   // hmiStns[1].wip[18].pnCode[6] := 1000;
   // hmiStns[1].wip[18].pnCode[7] := 1000;
   // hmiStns[1].wip[19].pnCode[0] := 1000;
   // hmiStns[1].wip[19].pnCode[1] := 1000;
   // hmiStns[1].wip[19].pnCode[2] := 1000;
   // hmiStns[1].wip[19].pnCode[3] := 1000;
   // hmiStns[1].wip[19].pnCode[4] := 1000;
   // hmiStns[1].wip[19].pnCode[5] := 1000;
   // hmiStns[1].wip[19].pnCode[6] := 1000;
   // hmiStns[1].wip[19].pnCode[7] := 1000;
   // hmiStns[1].wip[20].pnCode[0] := 1000;
   // hmiStns[1].wip[20].pnCode[1] := 1000;
   // hmiStns[1].wip[20].pnCode[2] := 1000;
   // hmiStns[1].wip[20].pnCode[3] := 1000;
   // hmiStns[1].wip[20].pnCode[4] := 1000;
   // hmiStns[1].wip[20].pnCode[5] := 1000;
   // hmiStns[1].wip[20].pnCode[6] := 1000;
   // hmiStns[1].wip[20].pnCode[7] := 1000;
   // hmiStns[1].wip[21].pnCode[0] := 1000;
   // hmiStns[1].wip[21].pnCode[1] := 1000;
   // hmiStns[1].wip[21].pnCode[2] := 1000;
   // hmiStns[1].wip[21].pnCode[3] := 1000;
   // hmiStns[1].wip[21].pnCode[4] := 1000;
   // hmiStns[1].wip[21].pnCode[5] := 1000;
   // hmiStns[1].wip[21].pnCode[6] := 1000;
   // hmiStns[1].wip[21].pnCode[7] := 1000;
   // hmiStns[1].wip[22].pnCode[0] := 1000;
   // hmiStns[1].wip[22].pnCode[1] := 1000;
   // hmiStns[1].wip[22].pnCode[2] := 1000;
   // hmiStns[1].wip[22].pnCode[3] := 1000;
   // hmiStns[1].wip[22].pnCode[4] := 1000;
   // hmiStns[1].wip[22].pnCode[5] := 1000;
   // hmiStns[1].wip[22].pnCode[6] := 1000;
   // hmiStns[1].wip[22].pnCode[7] := 1000;
   // hmiStns[1].wip[23].pnCode[0] := 1000;
   // hmiStns[1].wip[23].pnCode[1] := 1000;
   // hmiStns[1].wip[23].pnCode[2] := 1000;
   // hmiStns[1].wip[23].pnCode[3] := 1000;
   // hmiStns[1].wip[23].pnCode[4] := 1000;
   // hmiStns[1].wip[23].pnCode[5] := 1000;
   // hmiStns[1].wip[23].pnCode[6] := 1000;
   // hmiStns[1].wip[23].pnCode[7] := 1000;
   // hmiStns[1].wip[24].pnCode[0] := 1000;
   // hmiStns[1].wip[24].pnCode[1] := 1000;
   // hmiStns[1].wip[24].pnCode[2] := 1000;
   // hmiStns[1].wip[24].pnCode[3] := 1000;
   // hmiStns[1].wip[24].pnCode[4] := 1000;
   // hmiStns[1].wip[24].pnCode[5] := 1000;
   // hmiStns[1].wip[24].pnCode[6] := 1000;
   // hmiStns[1].wip[24].pnCode[7] := 1000;
   // hmiStns[1].wip[25].pnCode[0] := 1000;
   // hmiStns[1].wip[25].pnCode[1] := 1000;
   // hmiStns[1].wip[25].pnCode[2] := 1000;
   // hmiStns[1].wip[25].pnCode[3] := 1000;
   // hmiStns[1].wip[25].pnCode[4] := 1000;
   // hmiStns[1].wip[25].pnCode[5] := 1000;
   // hmiStns[1].wip[25].pnCode[6] := 1000;
   // hmiStns[1].wip[25].pnCode[7] := 1000;
   // hmiStns[1].wip[26].pnCode[0] := 1000;
   // hmiStns[1].wip[26].pnCode[1] := 1000;
   // hmiStns[1].wip[26].pnCode[2] := 1000;
   // hmiStns[1].wip[26].pnCode[3] := 1000;
   // hmiStns[1].wip[26].pnCode[4] := 1000;
   // hmiStns[1].wip[26].pnCode[5] := 1000;
   // hmiStns[1].wip[26].pnCode[6] := 1000;
   // hmiStns[1].wip[26].pnCode[7] := 1000;
   // hmiStns[1].wip[27].pnCode[0] := 1000;
   // hmiStns[1].wip[27].pnCode[1] := 1000;
   // hmiStns[1].wip[27].pnCode[2] := 1000;
   // hmiStns[1].wip[27].pnCode[3] := 1000;
   // hmiStns[1].wip[27].pnCode[4] := 1000;
   // hmiStns[1].wip[27].pnCode[5] := 1000;
   // hmiStns[1].wip[27].pnCode[6] := 1000;
   // hmiStns[1].wip[27].pnCode[7] := 1000;
   // hmiStns[1].wip[28].pnCode[0] := 1000;
   // hmiStns[1].wip[28].pnCode[1] := 1000;
   // hmiStns[1].wip[28].pnCode[2] := 1000;
   // hmiStns[1].wip[28].pnCode[3] := 1000;
   // hmiStns[1].wip[28].pnCode[4] := 1000;
   // hmiStns[1].wip[28].pnCode[5] := 1000;
   // hmiStns[1].wip[28].pnCode[6] := 1000;
   // hmiStns[1].wip[28].pnCode[7] := 1000;
   // hmiStns[1].wip[29].pnCode[0] := 1000;
   // hmiStns[1].wip[29].pnCode[1] := 1000;
   // hmiStns[1].wip[29].pnCode[2] := 1000;
   // hmiStns[1].wip[29].pnCode[3] := 1000;
   // hmiStns[1].wip[29].pnCode[4] := 1000;
   // hmiStns[1].wip[29].pnCode[5] := 1000;
   // hmiStns[1].wip[29].pnCode[6] := 1000;
   // hmiStns[1].wip[29].pnCode[7] := 1000;
   // hmiStns[1].wip[30].pnCode[0] := 1000;
   // hmiStns[1].wip[30].pnCode[1] := 1000;
   // hmiStns[1].wip[30].pnCode[2] := 1000;
   // hmiStns[1].wip[30].pnCode[3] := 1000;
   // hmiStns[1].wip[30].pnCode[4] := 1000;
   // hmiStns[1].wip[30].pnCode[5] := 1000;
   // hmiStns[1].wip[30].pnCode[6] := 1000;
   // hmiStns[1].wip[30].pnCode[7] := 1000;
   // hmiStns[1].wip[31].pnCode[0] := 1000;
   // hmiStns[1].wip[31].pnCode[1] := 1000;
   // hmiStns[1].wip[31].pnCode[2] := 1000;
   // hmiStns[1].wip[31].pnCode[3] := 1000;
   // hmiStns[1].wip[31].pnCode[4] := 1000;
   // hmiStns[1].wip[31].pnCode[5] := 1000;
   // hmiStns[1].wip[31].pnCode[6] := 1000;
   // hmiStns[1].wip[31].pnCode[7] := 1000;
   // hmiStns[1].wip[32].pnCode[0] := 1000;
   // hmiStns[1].wip[32].pnCode[1] := 1000;
   // hmiStns[1].wip[32].pnCode[2] := 1000;
   // hmiStns[1].wip[32].pnCode[3] := 1000;
   // hmiStns[1].wip[32].pnCode[4] := 1000;
   // hmiStns[1].wip[32].pnCode[5] := 1000;
   // hmiStns[1].wip[32].pnCode[6] := 1000;
   // hmiStns[1].wip[32].pnCode[7] := 1000;
   // hmiStns[1].wip[33].pnCode[0] := 1000;
   // hmiStns[1].wip[33].pnCode[1] := 1000;
   // hmiStns[1].wip[33].pnCode[2] := 1000;
   // hmiStns[1].wip[33].pnCode[3] := 1000;
   // hmiStns[1].wip[33].pnCode[4] := 1000;
   // hmiStns[1].wip[33].pnCode[5] := 1000;
   // hmiStns[1].wip[33].pnCode[6] := 1000;
   // hmiStns[1].wip[33].pnCode[7] := 1000;
   // hmiStns[1].wip[34].pnCode[0] := 1000;
   // hmiStns[1].wip[34].pnCode[1] := 1000;
   // hmiStns[1].wip[34].pnCode[2] := 1000;
   // hmiStns[1].wip[34].pnCode[3] := 1000;
   // hmiStns[1].wip[34].pnCode[4] := 1000;
   // hmiStns[1].wip[34].pnCode[5] := 1000;
   // hmiStns[1].wip[34].pnCode[6] := 1000;
   // hmiStns[1].wip[34].pnCode[7] := 1000;
   // hmiStns[1].wip[35].pnCode[0] := 1000;
   // hmiStns[1].wip[35].pnCode[1] := 1000;
   // hmiStns[1].wip[35].pnCode[2] := 1000;
   // hmiStns[1].wip[35].pnCode[3] := 1000;
   // hmiStns[1].wip[35].pnCode[4] := 1000;
   // hmiStns[1].wip[35].pnCode[5] := 1000;
   // hmiStns[1].wip[35].pnCode[6] := 1000;
   // hmiStns[1].wip[35].pnCode[7] := 1000;
   // hmiStns[1].wip[36].pnCode[0] := 1000;
   // hmiStns[1].wip[36].pnCode[1] := 1000;
   // hmiStns[1].wip[36].pnCode[2] := 1000;
   // hmiStns[1].wip[36].pnCode[3] := 1000;
   // hmiStns[1].wip[36].pnCode[4] := 1000;
   // hmiStns[1].wip[36].pnCode[5] := 1000;
   // hmiStns[1].wip[36].pnCode[6] := 1000;
   // hmiStns[1].wip[36].pnCode[7] := 1000;
   // hmiStns[1].wip[37].pnCode[0] := 1000;
   // hmiStns[1].wip[37].pnCode[1] := 1000;
   // hmiStns[1].wip[37].pnCode[2] := 1000;
   // hmiStns[1].wip[37].pnCode[3] := 1000;
   // hmiStns[1].wip[37].pnCode[4] := 1000;
   // hmiStns[1].wip[37].pnCode[5] := 1000;
   // hmiStns[1].wip[37].pnCode[6] := 1000;
   // hmiStns[1].wip[37].pnCode[7] := 1000;
   // hmiStns[1].wip[38].pnCode[0] := 1000;
   // hmiStns[1].wip[38].pnCode[1] := 1000;
   // hmiStns[1].wip[38].pnCode[2] := 1000;
   // hmiStns[1].wip[38].pnCode[3] := 1000;
   // hmiStns[1].wip[38].pnCode[4] := 1000;
   // hmiStns[1].wip[38].pnCode[5] := 1000;
   // hmiStns[1].wip[38].pnCode[6] := 1000;
   // hmiStns[1].wip[38].pnCode[7] := 1000;
   // hmiStns[1].wip[39].pnCode[0] := 1000;
   // hmiStns[1].wip[39].pnCode[1] := 1000;
   // hmiStns[1].wip[39].pnCode[2] := 1000;
   // hmiStns[1].wip[39].pnCode[3] := 1000;
   // hmiStns[1].wip[39].pnCode[4] := 1000;
   // hmiStns[1].wip[39].pnCode[5] := 1000;
   // hmiStns[1].wip[39].pnCode[6] := 1000;
   // hmiStns[1].wip[39].pnCode[7] := 1000;
   // hmiStns[1].wip[40].pnCode[0] := 1000;
   // hmiStns[1].wip[40].pnCode[1] := 1000;
   // hmiStns[1].wip[40].pnCode[2] := 1000;
   // hmiStns[1].wip[40].pnCode[3] := 1000;
   // hmiStns[1].wip[40].pnCode[4] := 1000;
   // hmiStns[1].wip[40].pnCode[5] := 1000;
   // hmiStns[1].wip[40].pnCode[6] := 1000;
   // hmiStns[1].wip[40].pnCode[7] := 1000;
   // hmiStns[1].wip[41].pnCode[0] := 1000;
   // hmiStns[1].wip[41].pnCode[1] := 1000;
   // hmiStns[1].wip[41].pnCode[2] := 1000;
   // hmiStns[1].wip[41].pnCode[3] := 1000;
   // hmiStns[1].wip[41].pnCode[4] := 1000;
   // hmiStns[1].wip[41].pnCode[5] := 1000;
   // hmiStns[1].wip[41].pnCode[6] := 1000;
   // hmiStns[1].wip[41].pnCode[7] := 1000;
   // hmiStns[1].wip[42].pnCode[0] := 1000;
   // hmiStns[1].wip[42].pnCode[1] := 1000;
   // hmiStns[1].wip[42].pnCode[2] := 1000;
   // hmiStns[1].wip[42].pnCode[3] := 1000;
   // hmiStns[1].wip[42].pnCode[4] := 1000;
   // hmiStns[1].wip[42].pnCode[5] := 1000;
   // hmiStns[1].wip[42].pnCode[6] := 1000;
   // hmiStns[1].wip[42].pnCode[7] := 1000;
   // hmiStns[1].wip[43].pnCode[0] := 1000;
   // hmiStns[1].wip[43].pnCode[1] := 1000;
   // hmiStns[1].wip[43].pnCode[2] := 1000;
   // hmiStns[1].wip[43].pnCode[3] := 1000;
   // hmiStns[1].wip[43].pnCode[4] := 1000;
   // hmiStns[1].wip[43].pnCode[5] := 1000;
   // hmiStns[1].wip[43].pnCode[6] := 1000;
   // hmiStns[1].wip[43].pnCode[7] := 1000;
   // hmiStns[1].wip[44].pnCode[0] := 1000;
   // hmiStns[1].wip[44].pnCode[1] := 1000;
   // hmiStns[1].wip[44].pnCode[2] := 1000;
   // hmiStns[1].wip[44].pnCode[3] := 1000;
   // hmiStns[1].wip[44].pnCode[4] := 1000;
   // hmiStns[1].wip[44].pnCode[5] := 1000;
   // hmiStns[1].wip[44].pnCode[6] := 1000;
   // hmiStns[1].wip[44].pnCode[7] := 1000;
   // hmiStns[1].wip[45].pnCode[0] := 1000;
   // hmiStns[1].wip[45].pnCode[1] := 1000;
   // hmiStns[1].wip[45].pnCode[2] := 1000;
   // hmiStns[1].wip[45].pnCode[3] := 1000;
   // hmiStns[1].wip[45].pnCode[4] := 1000;
   // hmiStns[1].wip[45].pnCode[5] := 1000;
   // hmiStns[1].wip[45].pnCode[6] := 1000;
   // hmiStns[1].wip[45].pnCode[7] := 1000;
   // hmiStns[1].wip[46].pnCode[0] := 1000;
   // hmiStns[1].wip[46].pnCode[1] := 1000;
   // hmiStns[1].wip[46].pnCode[2] := 1000;
   // hmiStns[1].wip[46].pnCode[3] := 1000;
   // hmiStns[1].wip[46].pnCode[4] := 1000;
   // hmiStns[1].wip[46].pnCode[5] := 1000;
   // hmiStns[1].wip[46].pnCode[6] := 1000;
   // hmiStns[1].wip[46].pnCode[7] := 1000;
   // hmiStns[1].wip[47].pnCode[0] := 1000;
   // hmiStns[1].wip[47].pnCode[1] := 1000;
   // hmiStns[1].wip[47].pnCode[2] := 1000;
   // hmiStns[1].wip[47].pnCode[3] := 1000;
   // hmiStns[1].wip[47].pnCode[4] := 1000;
   // hmiStns[1].wip[47].pnCode[5] := 1000;
   // hmiStns[1].wip[47].pnCode[6] := 1000;
   // hmiStns[1].wip[47].pnCode[7] := 1000;
   // hmiStns[1].wip[48].pnCode[0] := 1000;
   // hmiStns[1].wip[48].pnCode[1] := 1000;
   // hmiStns[1].wip[48].pnCode[2] := 1000;
   // hmiStns[1].wip[48].pnCode[3] := 1000;
   // hmiStns[1].wip[48].pnCode[4] := 1000;
   // hmiStns[1].wip[48].pnCode[5] := 1000;
   // hmiStns[1].wip[48].pnCode[6] := 1000;
   // hmiStns[1].wip[48].pnCode[7] := 1000;
   // hmiStns[1].wip[49].pnCode[0] := 1000;
   // hmiStns[1].wip[49].pnCode[1] := 1000;
   // hmiStns[1].wip[49].pnCode[2] := 1000;
   // hmiStns[1].wip[49].pnCode[3] := 1000;
   // hmiStns[1].wip[49].pnCode[4] := 1000;
   // hmiStns[1].wip[49].pnCode[5] := 1000;
   // hmiStns[1].wip[49].pnCode[6] := 1000;
   // hmiStns[1].wip[49].pnCode[7] := 1000;
   // hmiStns[2].pStn := 27;
   // hmiStns[2].wip[0].pnCode[0] := 1000;
   // hmiStns[2].wip[0].pnCode[1] := 244000;
   // hmiStns[2].wip[0].pnCode[2] := 149000;
   // hmiStns[2].wip[0].pnCode[3] := 1000;
   // hmiStns[2].wip[0].pnCode[4] := 1000;
   // hmiStns[2].wip[0].pnCode[5] := 1000;
   // hmiStns[2].wip[0].pnCode[6] := 148000;
   // hmiStns[2].wip[0].pnCode[7] := 150000;
   // hmiStns[2].wip[1].pnCode[0] := 1000;
   // hmiStns[2].wip[1].pnCode[1] := 244000;
   // hmiStns[2].wip[1].pnCode[2] := 54000;
   // hmiStns[2].wip[1].pnCode[3] := 1000;
   // hmiStns[2].wip[1].pnCode[4] := 1000;
   // hmiStns[2].wip[1].pnCode[5] := 1000;
   // hmiStns[2].wip[1].pnCode[6] := 32000;
   // hmiStns[2].wip[1].pnCode[7] := 72000;
   // hmiStns[2].wip[2].pnCode[0] := 1000;
   // hmiStns[2].wip[2].pnCode[1] := 244000;
   // hmiStns[2].wip[2].pnCode[2] := 58000;
   // hmiStns[2].wip[2].pnCode[3] := 1000;
   // hmiStns[2].wip[2].pnCode[4] := 1000;
   // hmiStns[2].wip[2].pnCode[5] := 1000;
   // hmiStns[2].wip[2].pnCode[6] := 26000;
   // hmiStns[2].wip[2].pnCode[7] := 19000;
   // hmiStns[2].wip[3].pnCode[0] := 1000;
   // hmiStns[2].wip[3].pnCode[1] := 244000;
   // hmiStns[2].wip[3].pnCode[2] := 85000;
   // hmiStns[2].wip[3].pnCode[3] := 1000;
   // hmiStns[2].wip[3].pnCode[4] := 1000;
   // hmiStns[2].wip[3].pnCode[5] := 1000;
   // hmiStns[2].wip[3].pnCode[6] := 32000;
   // hmiStns[2].wip[3].pnCode[7] := 72000;
   // hmiStns[2].wip[4].pnCode[0] := 1000;
   // hmiStns[2].wip[4].pnCode[1] := 244000;
   // hmiStns[2].wip[4].pnCode[2] := 71000;
   // hmiStns[2].wip[4].pnCode[3] := 73000;
   // hmiStns[2].wip[4].pnCode[4] := 1000;
   // hmiStns[2].wip[4].pnCode[5] := 59000;
   // hmiStns[2].wip[4].pnCode[6] := 34000;
   // hmiStns[2].wip[4].pnCode[7] := 74000;
   // hmiStns[2].wip[5].pnCode[0] := 1000;
   // hmiStns[2].wip[5].pnCode[1] := 244000;
   // hmiStns[2].wip[5].pnCode[2] := 128000;
   // hmiStns[2].wip[5].pnCode[3] := 1000;
   // hmiStns[2].wip[5].pnCode[4] := 1000;
   // hmiStns[2].wip[5].pnCode[5] := 101000;
   // hmiStns[2].wip[5].pnCode[6] := 102000;
   // hmiStns[2].wip[5].pnCode[7] := 129000;
   // hmiStns[2].wip[6].pnCode[0] := 1000;
   // hmiStns[2].wip[6].pnCode[1] := 244000;
   // hmiStns[2].wip[6].pnCode[2] := 123000;
   // hmiStns[2].wip[6].pnCode[3] := 124000;
   // hmiStns[2].wip[6].pnCode[4] := 1000;
   // hmiStns[2].wip[6].pnCode[5] := 103000;
   // hmiStns[2].wip[6].pnCode[6] := 104000;
   // hmiStns[2].wip[6].pnCode[7] := 134000;
   // hmiStns[2].wip[7].pnCode[0] := 1000;
   // hmiStns[2].wip[7].pnCode[1] := 244000;
   // hmiStns[2].wip[7].pnCode[2] := 101000;
   // hmiStns[2].wip[7].pnCode[3] := 129000;
   // hmiStns[2].wip[7].pnCode[4] := 1000;
   // hmiStns[2].wip[7].pnCode[5] := 103000;
   // hmiStns[2].wip[7].pnCode[6] := 105000;
   // hmiStns[2].wip[7].pnCode[7] := 134000;
   // hmiStns[2].wip[8].pnCode[0] := 1000;
   // hmiStns[2].wip[8].pnCode[1] := 244000;
   // hmiStns[2].wip[8].pnCode[2] := 106000;
   // hmiStns[2].wip[8].pnCode[3] := 124000;
   // hmiStns[2].wip[8].pnCode[4] := 1000;
   // hmiStns[2].wip[8].pnCode[5] := 107000;
   // hmiStns[2].wip[8].pnCode[6] := 108000;
   // hmiStns[2].wip[8].pnCode[7] := 134000;
   // hmiStns[2].wip[9].pnCode[0] := 1000;
   // hmiStns[2].wip[9].pnCode[1] := 244000;
   // hmiStns[2].wip[9].pnCode[2] := 101000;
   // hmiStns[2].wip[9].pnCode[3] := 1000;
   // hmiStns[2].wip[9].pnCode[4] := 1000;
   // hmiStns[2].wip[9].pnCode[5] := 128000;
   // hmiStns[2].wip[9].pnCode[6] := 108000;
   // hmiStns[2].wip[9].pnCode[7] := 129000;
   // hmiStns[2].wip[10].pnCode[0] := 1000;
   // hmiStns[2].wip[10].pnCode[1] := 244000;
   // hmiStns[2].wip[10].pnCode[2] := 101000;
   // hmiStns[2].wip[10].pnCode[3] := 129000;
   // hmiStns[2].wip[10].pnCode[4] := 1000;
   // hmiStns[2].wip[10].pnCode[5] := 107000;
   // hmiStns[2].wip[10].pnCode[6] := 108000;
   // hmiStns[2].wip[10].pnCode[7] := 124000;
   // hmiStns[2].wip[11].pnCode[0] := 1000;
   // hmiStns[2].wip[11].pnCode[1] := 244000;
   // hmiStns[2].wip[11].pnCode[2] := 109000;
   // hmiStns[2].wip[11].pnCode[3] := 1000;
   // hmiStns[2].wip[11].pnCode[4] := 1000;
   // hmiStns[2].wip[11].pnCode[5] := 1000;
   // hmiStns[2].wip[11].pnCode[6] := 108000;
   // hmiStns[2].wip[11].pnCode[7] := 110000;
   // hmiStns[2].wip[12].pnCode[0] := 1000;
   // hmiStns[2].wip[12].pnCode[1] := 244000;
   // hmiStns[2].wip[12].pnCode[2] := 111000;
   // hmiStns[2].wip[12].pnCode[3] := 114000;
   // hmiStns[2].wip[12].pnCode[4] := 1000;
   // hmiStns[2].wip[12].pnCode[5] := 113000;
   // hmiStns[2].wip[12].pnCode[6] := 115000;
   // hmiStns[2].wip[12].pnCode[7] := 112000;
   // hmiStns[2].wip[13].pnCode[0] := 1000;
   // hmiStns[2].wip[13].pnCode[1] := 244000;
   // hmiStns[2].wip[13].pnCode[2] := 116000;
   // hmiStns[2].wip[13].pnCode[3] := 1000;
   // hmiStns[2].wip[13].pnCode[4] := 1000;
   // hmiStns[2].wip[13].pnCode[5] := 113000;
   // hmiStns[2].wip[13].pnCode[6] := 115000;
   // hmiStns[2].wip[13].pnCode[7] := 114000;
   // hmiStns[2].wip[14].pnCode[0] := 1000;
   // hmiStns[2].wip[14].pnCode[1] := 244000;
   // hmiStns[2].wip[14].pnCode[2] := 117000;
   // hmiStns[2].wip[14].pnCode[3] := 112000;
   // hmiStns[2].wip[14].pnCode[4] := 1000;
   // hmiStns[2].wip[14].pnCode[5] := 119000;
   // hmiStns[2].wip[14].pnCode[6] := 115000;
   // hmiStns[2].wip[14].pnCode[7] := 118000;
   // hmiStns[2].wip[15].pnCode[0] := 1000;
   // hmiStns[2].wip[15].pnCode[1] := 244000;
   // hmiStns[2].wip[15].pnCode[2] := 117000;
   // hmiStns[2].wip[15].pnCode[3] := 118000;
   // hmiStns[2].wip[15].pnCode[4] := 1000;
   // hmiStns[2].wip[15].pnCode[5] := 119000;
   // hmiStns[2].wip[15].pnCode[6] := 121000;
   // hmiStns[2].wip[15].pnCode[7] := 112000;
   // hmiStns[2].wip[16].pnCode[0] := 1000;
   // hmiStns[2].wip[16].pnCode[1] := 244000;
   // hmiStns[2].wip[16].pnCode[2] := 120000;
   // hmiStns[2].wip[16].pnCode[3] := 1000;
   // hmiStns[2].wip[16].pnCode[4] := 1000;
   // hmiStns[2].wip[16].pnCode[5] := 122000;
   // hmiStns[2].wip[16].pnCode[6] := 115000;
   // hmiStns[2].wip[16].pnCode[7] := 112000;
   // hmiStns[2].wip[17].pnCode[0] := 1000;
   // hmiStns[2].wip[17].pnCode[1] := 244000;
   // hmiStns[2].wip[17].pnCode[2] := 125000;
   // hmiStns[2].wip[17].pnCode[3] := 126000;
   // hmiStns[2].wip[17].pnCode[4] := 1000;
   // hmiStns[2].wip[17].pnCode[5] := 123000;
   // hmiStns[2].wip[17].pnCode[6] := 108000;
   // hmiStns[2].wip[17].pnCode[7] := 124000;
   // hmiStns[2].wip[18].pnCode[0] := 1000;
   // hmiStns[2].wip[18].pnCode[1] := 244000;
   // hmiStns[2].wip[18].pnCode[2] := 101000;
   // hmiStns[2].wip[18].pnCode[3] := 1000;
   // hmiStns[2].wip[18].pnCode[4] := 1000;
   // hmiStns[2].wip[18].pnCode[5] := 128000;
   // hmiStns[2].wip[18].pnCode[6] := 127000;
   // hmiStns[2].wip[18].pnCode[7] := 129000;
   // hmiStns[2].wip[19].pnCode[0] := 1000;
   // hmiStns[2].wip[19].pnCode[1] := 244000;
   // hmiStns[2].wip[19].pnCode[2] := 128000;
   // hmiStns[2].wip[19].pnCode[3] := 124000;
   // hmiStns[2].wip[19].pnCode[4] := 1000;
   // hmiStns[2].wip[19].pnCode[5] := 123000;
   // hmiStns[2].wip[19].pnCode[6] := 130000;
   // hmiStns[2].wip[19].pnCode[7] := 129000;
   // hmiStns[2].wip[20].pnCode[0] := 1000;
   // hmiStns[2].wip[20].pnCode[1] := 244000;
   // hmiStns[2].wip[20].pnCode[2] := 131000;
   // hmiStns[2].wip[20].pnCode[3] := 1000;
   // hmiStns[2].wip[20].pnCode[4] := 1000;
   // hmiStns[2].wip[20].pnCode[5] := 1000;
   // hmiStns[2].wip[20].pnCode[6] := 127000;
   // hmiStns[2].wip[20].pnCode[7] := 132000;
   // hmiStns[2].wip[21].pnCode[0] := 1000;
   // hmiStns[2].wip[21].pnCode[1] := 244000;
   // hmiStns[2].wip[21].pnCode[2] := 133000;
   // hmiStns[2].wip[21].pnCode[3] := 1000;
   // hmiStns[2].wip[21].pnCode[4] := 1000;
   // hmiStns[2].wip[21].pnCode[5] := 1000;
   // hmiStns[2].wip[21].pnCode[6] := 144000;
   // hmiStns[2].wip[21].pnCode[7] := 134000;
   // hmiStns[2].wip[22].pnCode[0] := 1000;
   // hmiStns[2].wip[22].pnCode[1] := 244000;
   // hmiStns[2].wip[22].pnCode[2] := 135000;
   // hmiStns[2].wip[22].pnCode[3] := 1000;
   // hmiStns[2].wip[22].pnCode[4] := 1000;
   // hmiStns[2].wip[22].pnCode[5] := 1000;
   // hmiStns[2].wip[22].pnCode[6] := 144000;
   // hmiStns[2].wip[22].pnCode[7] := 136000;
   // hmiStns[2].wip[23].pnCode[0] := 1000;
   // hmiStns[2].wip[23].pnCode[1] := 244000;
   // hmiStns[2].wip[23].pnCode[2] := 143000;
   // hmiStns[2].wip[23].pnCode[3] := 1000;
   // hmiStns[2].wip[23].pnCode[4] := 1000;
   // hmiStns[2].wip[23].pnCode[5] := 1000;
   // hmiStns[2].wip[23].pnCode[6] := 144000;
   // hmiStns[2].wip[23].pnCode[7] := 134000;
   // hmiStns[2].wip[24].pnCode[0] := 1000;
   // hmiStns[2].wip[24].pnCode[1] := 244000;
   // hmiStns[2].wip[24].pnCode[2] := 137000;
   // hmiStns[2].wip[24].pnCode[3] := 1000;
   // hmiStns[2].wip[24].pnCode[4] := 1000;
   // hmiStns[2].wip[24].pnCode[5] := 1000;
   // hmiStns[2].wip[24].pnCode[6] := 144000;
   // hmiStns[2].wip[24].pnCode[7] := 136000;
   // hmiStns[2].wip[25].pnCode[0] := 1000;
   // hmiStns[2].wip[25].pnCode[1] := 244000;
   // hmiStns[2].wip[25].pnCode[2] := 138000;
   // hmiStns[2].wip[25].pnCode[3] := 1000;
   // hmiStns[2].wip[25].pnCode[4] := 1000;
   // hmiStns[2].wip[25].pnCode[5] := 1000;
   // hmiStns[2].wip[25].pnCode[6] := 141000;
   // hmiStns[2].wip[25].pnCode[7] := 129000;
   // hmiStns[2].wip[26].pnCode[0] := 1000;
   // hmiStns[2].wip[26].pnCode[1] := 244000;
   // hmiStns[2].wip[26].pnCode[2] := 139000;
   // hmiStns[2].wip[26].pnCode[3] := 1000;
   // hmiStns[2].wip[26].pnCode[4] := 1000;
   // hmiStns[2].wip[26].pnCode[5] := 1000;
   // hmiStns[2].wip[26].pnCode[6] := 141000;
   // hmiStns[2].wip[26].pnCode[7] := 140000;
   // hmiStns[2].wip[27].pnCode[0] := 1000;
   // hmiStns[2].wip[27].pnCode[1] := 244000;
   // hmiStns[2].wip[27].pnCode[2] := 142000;
   // hmiStns[2].wip[27].pnCode[3] := 1000;
   // hmiStns[2].wip[27].pnCode[4] := 1000;
   // hmiStns[2].wip[27].pnCode[5] := 1000;
   // hmiStns[2].wip[27].pnCode[6] := 141000;
   // hmiStns[2].wip[27].pnCode[7] := 126000;
   // hmiStns[2].wip[28].pnCode[0] := 1000;
   // hmiStns[2].wip[28].pnCode[1] := 244000;
   // hmiStns[2].wip[28].pnCode[2] := 149000;
   // hmiStns[2].wip[28].pnCode[3] := 1000;
   // hmiStns[2].wip[28].pnCode[4] := 1000;
   // hmiStns[2].wip[28].pnCode[5] := 1000;
   // hmiStns[2].wip[28].pnCode[6] := 145000;
   // hmiStns[2].wip[28].pnCode[7] := 150000;
   // hmiStns[2].wip[29].pnCode[0] := 1000;
   // hmiStns[2].wip[29].pnCode[1] := 244000;
   // hmiStns[2].wip[29].pnCode[2] := 146000;
   // hmiStns[2].wip[29].pnCode[3] := 1000;
   // hmiStns[2].wip[29].pnCode[4] := 1000;
   // hmiStns[2].wip[29].pnCode[5] := 1000;
   // hmiStns[2].wip[29].pnCode[6] := 148000;
   // hmiStns[2].wip[29].pnCode[7] := 147000;
   // hmiStns[2].wip[30].pnCode[0] := 1000;
   // hmiStns[2].wip[30].pnCode[1] := 244000;
   // hmiStns[2].wip[30].pnCode[2] := 160000;
   // hmiStns[2].wip[30].pnCode[3] := 1000;
   // hmiStns[2].wip[30].pnCode[4] := 1000;
   // hmiStns[2].wip[30].pnCode[5] := 1000;
   // hmiStns[2].wip[30].pnCode[6] := 145000;
   // hmiStns[2].wip[30].pnCode[7] := 161000;
   // hmiStns[2].wip[31].pnCode[0] := 1000;
   // hmiStns[2].wip[31].pnCode[1] := 244000;
   // hmiStns[2].wip[31].pnCode[2] := 164000;
   // hmiStns[2].wip[31].pnCode[3] := 1000;
   // hmiStns[2].wip[31].pnCode[4] := 1000;
   // hmiStns[2].wip[31].pnCode[5] := 1000;
   // hmiStns[2].wip[31].pnCode[6] := 148000;
   // hmiStns[2].wip[31].pnCode[7] := 147000;
   // hmiStns[2].wip[32].pnCode[0] := 1000;
   // hmiStns[2].wip[32].pnCode[1] := 244000;
   // hmiStns[2].wip[32].pnCode[2] := 160000;
   // hmiStns[2].wip[32].pnCode[3] := 1000;
   // hmiStns[2].wip[32].pnCode[4] := 1000;
   // hmiStns[2].wip[32].pnCode[5] := 1000;
   // hmiStns[2].wip[32].pnCode[6] := 148000;
   // hmiStns[2].wip[32].pnCode[7] := 161000;
   // hmiStns[2].wip[33].pnCode[0] := 1000;
   // hmiStns[2].wip[33].pnCode[1] := 244000;
   // hmiStns[2].wip[33].pnCode[2] := 153000;
   // hmiStns[2].wip[33].pnCode[3] := 152000;
   // hmiStns[2].wip[33].pnCode[4] := 1000;
   // hmiStns[2].wip[33].pnCode[5] := 151000;
   // hmiStns[2].wip[33].pnCode[6] := 155000;
   // hmiStns[2].wip[33].pnCode[7] := 154000;
   // hmiStns[2].wip[34].pnCode[0] := 1000;
   // hmiStns[2].wip[34].pnCode[1] := 244000;
   // hmiStns[2].wip[34].pnCode[2] := 153000;
   // hmiStns[2].wip[34].pnCode[3] := 1000;
   // hmiStns[2].wip[34].pnCode[4] := 1000;
   // hmiStns[2].wip[34].pnCode[5] := 156000;
   // hmiStns[2].wip[34].pnCode[6] := 155000;
   // hmiStns[2].wip[34].pnCode[7] := 154000;
   // hmiStns[2].wip[35].pnCode[0] := 1000;
   // hmiStns[2].wip[35].pnCode[1] := 244000;
   // hmiStns[2].wip[35].pnCode[2] := 157000;
   // hmiStns[2].wip[35].pnCode[3] := 1000;
   // hmiStns[2].wip[35].pnCode[4] := 1000;
   // hmiStns[2].wip[35].pnCode[5] := 1000;
   // hmiStns[2].wip[35].pnCode[6] := 155000;
   // hmiStns[2].wip[35].pnCode[7] := 158000;
   // hmiStns[2].wip[36].pnCode[0] := 1000;
   // hmiStns[2].wip[36].pnCode[1] := 244000;
   // hmiStns[2].wip[36].pnCode[2] := 160000;
   // hmiStns[2].wip[36].pnCode[3] := 1000;
   // hmiStns[2].wip[36].pnCode[4] := 1000;
   // hmiStns[2].wip[36].pnCode[5] := 1000;
   // hmiStns[2].wip[36].pnCode[6] := 162000;
   // hmiStns[2].wip[36].pnCode[7] := 161000;
   // hmiStns[2].wip[37].pnCode[0] := 1000;
   // hmiStns[2].wip[37].pnCode[1] := 244000;
   // hmiStns[2].wip[37].pnCode[2] := 159000;
   // hmiStns[2].wip[37].pnCode[3] := 1000;
   // hmiStns[2].wip[37].pnCode[4] := 1000;
   // hmiStns[2].wip[37].pnCode[5] := 1000;
   // hmiStns[2].wip[37].pnCode[6] := 162000;
   // hmiStns[2].wip[37].pnCode[7] := 161000;
   // hmiStns[2].wip[38].pnCode[0] := 1000;
   // hmiStns[2].wip[38].pnCode[1] := 244000;
   // hmiStns[2].wip[38].pnCode[2] := 163000;
   // hmiStns[2].wip[38].pnCode[3] := 1000;
   // hmiStns[2].wip[38].pnCode[4] := 1000;
   // hmiStns[2].wip[38].pnCode[5] := 1000;
   // hmiStns[2].wip[38].pnCode[6] := 162000;
   // hmiStns[2].wip[38].pnCode[7] := 161000;
   // hmiStns[2].wip[39].pnCode[0] := 1000;
   // hmiStns[2].wip[39].pnCode[1] := 244000;
   // hmiStns[2].wip[39].pnCode[2] := 164000;
   // hmiStns[2].wip[39].pnCode[3] := 1000;
   // hmiStns[2].wip[39].pnCode[4] := 1000;
   // hmiStns[2].wip[39].pnCode[5] := 1000;
   // hmiStns[2].wip[39].pnCode[6] := 162000;
   // hmiStns[2].wip[39].pnCode[7] := 147000;
   // hmiStns[2].wip[40].pnCode[0] := 1000;
   // hmiStns[2].wip[40].pnCode[1] := 244000;
   // hmiStns[2].wip[40].pnCode[2] := 106000;
   // hmiStns[2].wip[40].pnCode[3] := 129000;
   // hmiStns[2].wip[40].pnCode[4] := 1000;
   // hmiStns[2].wip[40].pnCode[5] := 128000;
   // hmiStns[2].wip[40].pnCode[6] := 127000;
   // hmiStns[2].wip[40].pnCode[7] := 134000;
   // hmiStns[2].wip[41].pnCode[0] := 1000;
   // hmiStns[2].wip[41].pnCode[1] := 244000;
   // hmiStns[2].wip[41].pnCode[2] := 1000;
   // hmiStns[2].wip[41].pnCode[3] := 1000;
   // hmiStns[2].wip[41].pnCode[4] := 1000;
   // hmiStns[2].wip[41].pnCode[5] := 1000;
   // hmiStns[2].wip[41].pnCode[6] := 1000;
   // hmiStns[2].wip[41].pnCode[7] := 1000;
   // hmiStns[2].wip[42].pnCode[0] := 1000;
   // hmiStns[2].wip[42].pnCode[1] := 244000;
   // hmiStns[2].wip[42].pnCode[2] := 1000;
   // hmiStns[2].wip[42].pnCode[3] := 1000;
   // hmiStns[2].wip[42].pnCode[4] := 1000;
   // hmiStns[2].wip[42].pnCode[5] := 1000;
   // hmiStns[2].wip[42].pnCode[6] := 1000;
   // hmiStns[2].wip[42].pnCode[7] := 1000;
   // hmiStns[2].wip[43].pnCode[0] := 1000;
   // hmiStns[2].wip[43].pnCode[1] := 244000;
   // hmiStns[2].wip[43].pnCode[2] := 1000;
   // hmiStns[2].wip[43].pnCode[3] := 1000;
   // hmiStns[2].wip[43].pnCode[4] := 1000;
   // hmiStns[2].wip[43].pnCode[5] := 1000;
   // hmiStns[2].wip[43].pnCode[6] := 1000;
   // hmiStns[2].wip[43].pnCode[7] := 1000;
   // hmiStns[2].wip[44].pnCode[0] := 1000;
   // hmiStns[2].wip[44].pnCode[1] := 244000;
   // hmiStns[2].wip[44].pnCode[2] := 1000;
   // hmiStns[2].wip[44].pnCode[3] := 1000;
   // hmiStns[2].wip[44].pnCode[4] := 1000;
   // hmiStns[2].wip[44].pnCode[5] := 1000;
   // hmiStns[2].wip[44].pnCode[6] := 1000;
   // hmiStns[2].wip[44].pnCode[7] := 1000;
   // hmiStns[2].wip[45].pnCode[0] := 1000;
   // hmiStns[2].wip[45].pnCode[1] := 244000;
   // hmiStns[2].wip[45].pnCode[2] := 1000;
   // hmiStns[2].wip[45].pnCode[3] := 1000;
   // hmiStns[2].wip[45].pnCode[4] := 1000;
   // hmiStns[2].wip[45].pnCode[5] := 1000;
   // hmiStns[2].wip[45].pnCode[6] := 1000;
   // hmiStns[2].wip[45].pnCode[7] := 1000;
   // hmiStns[2].wip[46].pnCode[0] := 1000;
   // hmiStns[2].wip[46].pnCode[1] := 244000;
   // hmiStns[2].wip[46].pnCode[2] := 1000;
   // hmiStns[2].wip[46].pnCode[3] := 1000;
   // hmiStns[2].wip[46].pnCode[4] := 1000;
   // hmiStns[2].wip[46].pnCode[5] := 1000;
   // hmiStns[2].wip[46].pnCode[6] := 1000;
   // hmiStns[2].wip[46].pnCode[7] := 1000;
   // hmiStns[2].wip[47].pnCode[0] := 1000;
   // hmiStns[2].wip[47].pnCode[1] := 244000;
   // hmiStns[2].wip[47].pnCode[2] := 1000;
   // hmiStns[2].wip[47].pnCode[3] := 1000;
   // hmiStns[2].wip[47].pnCode[4] := 1000;
   // hmiStns[2].wip[47].pnCode[5] := 1000;
   // hmiStns[2].wip[47].pnCode[6] := 1000;
   // hmiStns[2].wip[47].pnCode[7] := 1000;
   // hmiStns[2].wip[48].pnCode[0] := 1000;
   // hmiStns[2].wip[48].pnCode[1] := 244000;
   // hmiStns[2].wip[48].pnCode[2] := 1000;
   // hmiStns[2].wip[48].pnCode[3] := 1000;
   // hmiStns[2].wip[48].pnCode[4] := 1000;
   // hmiStns[2].wip[48].pnCode[5] := 1000;
   // hmiStns[2].wip[48].pnCode[6] := 1000;
   // hmiStns[2].wip[48].pnCode[7] := 1000;
   // hmiStns[2].wip[49].pnCode[0] := 1000;
   // hmiStns[2].wip[49].pnCode[1] := 244000;
   // hmiStns[2].wip[49].pnCode[2] := 1000;
   // hmiStns[2].wip[49].pnCode[3] := 1000;
   // hmiStns[2].wip[49].pnCode[4] := 1000;
   // hmiStns[2].wip[49].pnCode[5] := 1000;
   // hmiStns[2].wip[49].pnCode[6] := 1000;
   // hmiStns[2].wip[49].pnCode[7] := 1000;
   // hmiStns[3].pStn := 28;
   // hmiStns[3].wip[0].pnCode[0] := 1000;
   // hmiStns[3].wip[0].pnCode[1] := 244000;
   // hmiStns[3].wip[0].pnCode[2] := 53000;
   // hmiStns[3].wip[0].pnCode[3] := 1000;
   // hmiStns[3].wip[0].pnCode[4] := 1000;
   // hmiStns[3].wip[0].pnCode[5] := 1000;
   // hmiStns[3].wip[0].pnCode[6] := 32000;
   // hmiStns[3].wip[0].pnCode[7] := 74000;
   // hmiStns[3].wip[1].pnCode[0] := 1000;
   // hmiStns[3].wip[1].pnCode[1] := 244000;
   // hmiStns[3].wip[1].pnCode[2] := 218000;
   // hmiStns[3].wip[1].pnCode[3] := 1000;
   // hmiStns[3].wip[1].pnCode[4] := 1000;
   // hmiStns[3].wip[1].pnCode[5] := 1000;
   // hmiStns[3].wip[1].pnCode[6] := 219000;
   // hmiStns[3].wip[1].pnCode[7] := 224000;
   // hmiStns[3].wip[2].pnCode[0] := 1000;
   // hmiStns[3].wip[2].pnCode[1] := 244000;
   // hmiStns[3].wip[2].pnCode[2] := 229000;
   // hmiStns[3].wip[2].pnCode[3] := 232000;
   // hmiStns[3].wip[2].pnCode[4] := 1000;
   // hmiStns[3].wip[2].pnCode[5] := 230000;
   // hmiStns[3].wip[2].pnCode[6] := 228000;
   // hmiStns[3].wip[2].pnCode[7] := 231000;
   // hmiStns[3].wip[3].pnCode[0] := 1000;
   // hmiStns[3].wip[3].pnCode[1] := 244000;
   // hmiStns[3].wip[3].pnCode[2] := 165000;
   // hmiStns[3].wip[3].pnCode[3] := 1000;
   // hmiStns[3].wip[3].pnCode[4] := 1000;
   // hmiStns[3].wip[3].pnCode[5] := 166000;
   // hmiStns[3].wip[3].pnCode[6] := 203000;
   // hmiStns[3].wip[3].pnCode[7] := 204000;
   // hmiStns[3].wip[4].pnCode[0] := 1000;
   // hmiStns[3].wip[4].pnCode[1] := 244000;
   // hmiStns[3].wip[4].pnCode[2] := 201000;
   // hmiStns[3].wip[4].pnCode[3] := 1000;
   // hmiStns[3].wip[4].pnCode[4] := 1000;
   // hmiStns[3].wip[4].pnCode[5] := 202000;
   // hmiStns[3].wip[4].pnCode[6] := 203000;
   // hmiStns[3].wip[4].pnCode[7] := 204000;
   // hmiStns[3].wip[5].pnCode[0] := 1000;
   // hmiStns[3].wip[5].pnCode[1] := 244000;
   // hmiStns[3].wip[5].pnCode[2] := 165000;
   // hmiStns[3].wip[5].pnCode[3] := 1000;
   // hmiStns[3].wip[5].pnCode[4] := 1000;
   // hmiStns[3].wip[5].pnCode[5] := 166000;
   // hmiStns[3].wip[5].pnCode[6] := 203000;
   // hmiStns[3].wip[5].pnCode[7] := 204000;
   // hmiStns[3].wip[6].pnCode[0] := 1000;
   // hmiStns[3].wip[6].pnCode[1] := 244000;
   // hmiStns[3].wip[6].pnCode[2] := 1000;
   // hmiStns[3].wip[6].pnCode[3] := 186000;
   // hmiStns[3].wip[6].pnCode[4] := 1000;
   // hmiStns[3].wip[6].pnCode[5] := 1000;
   // hmiStns[3].wip[6].pnCode[6] := 198000;
   // hmiStns[3].wip[6].pnCode[7] := 180000;
   // hmiStns[3].wip[7].pnCode[0] := 1000;
   // hmiStns[3].wip[7].pnCode[1] := 244000;
   // hmiStns[3].wip[7].pnCode[2] := 1000;
   // hmiStns[3].wip[7].pnCode[3] := 200000;
   // hmiStns[3].wip[7].pnCode[4] := 1000;
   // hmiStns[3].wip[7].pnCode[5] := 1000;
   // hmiStns[3].wip[7].pnCode[6] := 199000;
   // hmiStns[3].wip[7].pnCode[7] := 179000;
   // hmiStns[3].wip[8].pnCode[0] := 1000;
   // hmiStns[3].wip[8].pnCode[1] := 1000;
   // hmiStns[3].wip[8].pnCode[2] := 1000;
   // hmiStns[3].wip[8].pnCode[3] := 1000;
   // hmiStns[3].wip[8].pnCode[4] := 1000;
   // hmiStns[3].wip[8].pnCode[5] := 1000;
   // hmiStns[3].wip[8].pnCode[6] := 1000;
   // hmiStns[3].wip[8].pnCode[7] := 1000;
   // hmiStns[3].wip[9].pnCode[0] := 1000;
   // hmiStns[3].wip[9].pnCode[1] := 1000;
   // hmiStns[3].wip[9].pnCode[2] := 1000;
   // hmiStns[3].wip[9].pnCode[3] := 1000;
   // hmiStns[3].wip[9].pnCode[4] := 1000;
   // hmiStns[3].wip[9].pnCode[5] := 1000;
   // hmiStns[3].wip[9].pnCode[6] := 1000;
   // hmiStns[3].wip[9].pnCode[7] := 1000;
   // hmiStns[3].wip[10].pnCode[0] := 1000;
   // hmiStns[3].wip[10].pnCode[1] := 1000;
   // hmiStns[3].wip[10].pnCode[2] := 1000;
   // hmiStns[3].wip[10].pnCode[3] := 1000;
   // hmiStns[3].wip[10].pnCode[4] := 1000;
   // hmiStns[3].wip[10].pnCode[5] := 1000;
   // hmiStns[3].wip[10].pnCode[6] := 1000;
   // hmiStns[3].wip[10].pnCode[7] := 1000;
   // hmiStns[3].wip[11].pnCode[0] := 1000;
   // hmiStns[3].wip[11].pnCode[1] := 1000;
   // hmiStns[3].wip[11].pnCode[2] := 1000;
   // hmiStns[3].wip[11].pnCode[3] := 1000;
   // hmiStns[3].wip[11].pnCode[4] := 1000;
   // hmiStns[3].wip[11].pnCode[5] := 1000;
   // hmiStns[3].wip[11].pnCode[6] := 1000;
   // hmiStns[3].wip[11].pnCode[7] := 1000;
   // hmiStns[3].wip[12].pnCode[0] := 1000;
   // hmiStns[3].wip[12].pnCode[1] := 1000;